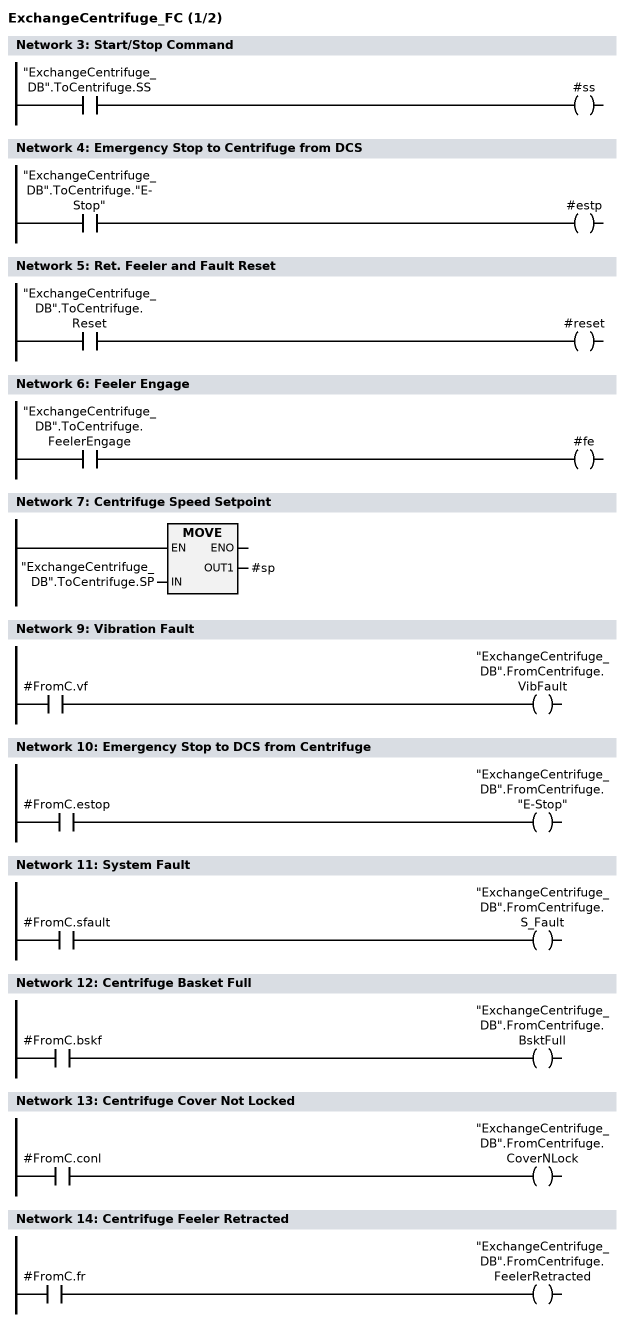
   RUNG wire#powerrail
      Contact( "ExchangeCentrifuge_DB".ToCentrifuge.SS )
      Coil( #ss )
   END_RUNG
   // the same network as SCL:
   #ss := "ExchangeCentrifuge_DB".ToCentrifuge.SS;
END_REGION

REGION Network 4: Emergency Stop to Centrifuge from DCS
   RUNG wire#powerrail
      Contact( "ExchangeCentrifuge_DB".ToCentrifuge."E-Stop" )
      Coil( #estp )
   END_RUNG
   // the same network as SCL:
   #estp := "ExchangeCentrifuge_DB".ToCentrifuge."E-Stop";
END_REGION

REGION Network 5: Ret. Feeler and Fault Reset
   RUNG wire#powerrail
      Contact( "ExchangeCentrifuge_DB".ToCentrifuge.Reset )
      Coil( #reset )
   END_RUNG
   // the same network as SCL:
   #reset := "ExchangeCentrifuge_DB".ToCentrifuge.Reset;
END_REGION

REGION Network 6: Feeler Engage
   RUNG wire#powerrail
      Contact( "ExchangeCentrifuge_DB".ToCentrifuge.FeelerEngage )
      Coil( #fe )
   END_RUNG
   // the same network as SCL:
   #fe := "ExchangeCentrifuge_DB".ToCentrifuge.FeelerEngage;
END_REGION

REGION Network 7: Centrifuge Speed Setpoint
   RUNG wire#powerrail
      Move(in := "ExchangeCentrifuge_DB".ToCentrifuge.SP, out1 => #sp)
   END_RUNG
   // the same network as SCL:
   #sp := "ExchangeCentrifuge_DB".ToCentrifuge.SP;
END_REGION

REGION Network 8: ////*********From Centrifuge to DCS**********////
   // Periphery Signal will be added to the contacts
END_REGION

REGION Network 9: Vibration Fault
   RUNG wire#powerrail
      Contact( #FromC.vf )
      Coil( "ExchangeCentrifuge_DB".FromCentrifuge.VibFault )
   END_RUNG
   // the same network as SCL:
   "ExchangeCentrifuge_DB".FromCentrifuge.VibFault := #FromC.vf;
END_REGION

REGION Network 10: Emergency Stop to DCS from Centrifuge
   RUNG wire#powerrail
      Contact( #FromC.estop )
      Coil( "ExchangeCentrifuge_DB".FromCentrifuge."E-Stop" )
   END_RUNG
   // the same network as SCL:
   "ExchangeCentrifuge_DB".FromCentrifuge."E-Stop" := #FromC.estop;
END_REGION

REGION Network 11: System Fault
   RUNG wire#powerrail
      Contact( #FromC.sfault )
      Coil( "ExchangeCentrifuge_DB".FromCentrifuge.S_Fault )
   END_RUNG
   // the same network as SCL:
   "ExchangeCentrifuge_DB".FromCentrifuge.S_Fault := #FromC.sfault;
END_REGION

REGION Network 12: Centrifuge Basket Full
   RUNG wire#powerrail
      Contact( #FromC.bskf )
      Coil( "ExchangeCentrifuge_DB".FromCentrifuge.BsktFull )
   END_RUNG
   // the same network as SCL:
   "ExchangeCentrifuge_DB".FromCentrifuge.BsktFull := #FromC.bskf;
END_REGION

REGION Network 13: Centrifuge Cover Not Locked
   RUNG wire#powerrail
      Contact( #FromC.conl )
      Coil( "ExchangeCentrifuge_DB".FromCentrifuge.CoverNLock )
   END_RUNG
   // the same network as SCL:
   "ExchangeCentrifuge_DB".FromCentrifuge.CoverNLock := #FromC.conl;
END_REGION

REGION Network 14: Centrifuge Feeler Retracted
   RUNG wire#powerrail
      Contact( #FromC.fr )
      Coil( "ExchangeCentrifuge_DB".FromCentrifuge.FeelerRetracted )
   END_RUNG
   // the same network as SCL:
   "ExchangeCentrifuge_DB".FromCentrifuge.FeelerRetracted := #FromC.fr;
END_REGION

REGION Network 15: Vibration Transmitter
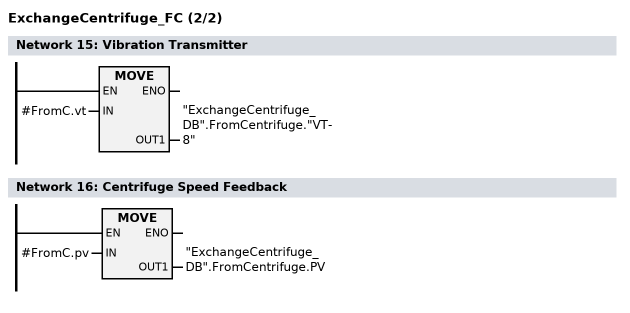
   RUNG wire#powerrail
      Move(in := #FromC.vt, out1 => "ExchangeCentrifuge_DB".FromCentrifuge."VT-8")
   END_RUNG
   // the same network as SCL:
   "ExchangeCentrifuge_DB".FromCentrifuge."VT-8" := #FromC.vt;
END_REGION

REGION Network 16: Centrifuge Speed Feedback
   RUNG wire#powerrail
      Move(in := #FromC.pv, out1 => "ExchangeCentrifuge_DB".FromCentrifuge.PV)
   END_RUNG
   // the same network as SCL:
   "ExchangeCentrifuge_DB".FromCentrifuge.PV := #FromC.pv;
END_REGION
END_FUNCTION

// folder: Outside Comms/ModBus Comms/CO/CO2/O2 R-401 Analizer

FUNCTION "Analizer_Modbus" : Void   // FC113, LAD
{ S7_Optimized_Access := 'TRUE' }
VERSION : 0.1
BEGIN

REGION Network 1: CO/CO2/O2 Analizer up to R-401 (Calcination)
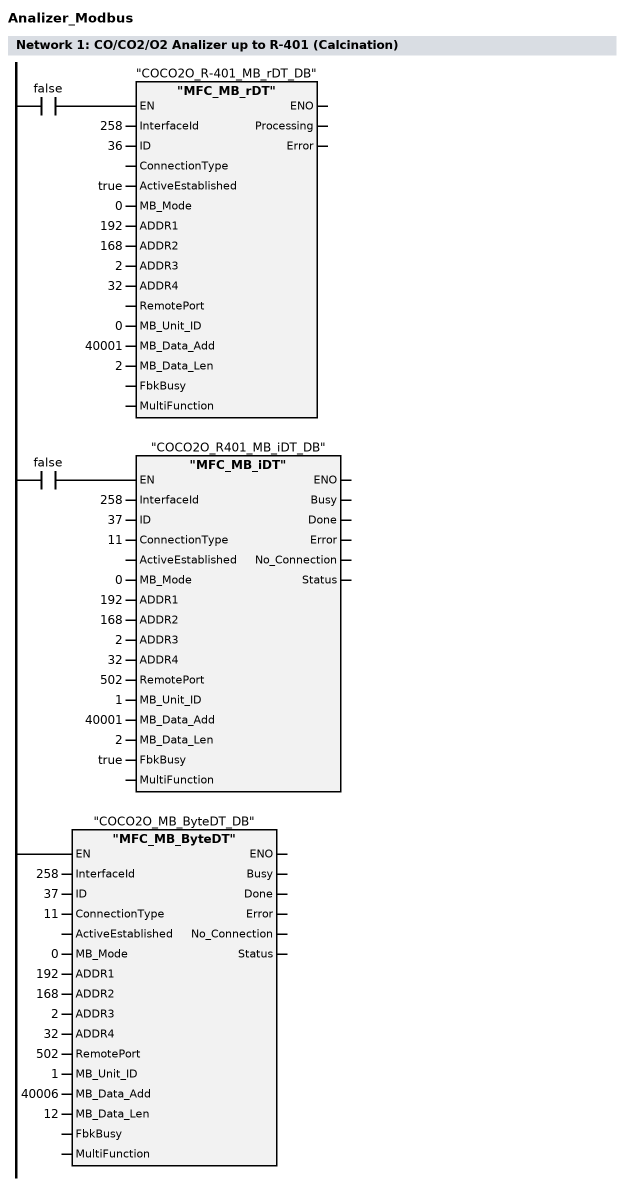
   RUNG wire#powerrail
      Contact( false )
      "COCO2O_R-401_MB_rDT_DB"(InterfaceId := 258, ID := 36, ConnectionType :=, ActiveEstablished := true, MB_Mode := 0, ADDR1 := 192, ADDR2 := 168, ADDR3 := 2, ADDR4 := 32, RemotePort :=, MB_Unit_ID := 0, MB_Data_Add := 40001, MB_Data_Len := 2, FbkBusy :=, MultiFunction :=, Processing =>, Error =>)
   END_RUNG
   RUNG wire#powerrail
      Contact( false )
      "COCO2O_R401_MB_iDT_DB"(InterfaceId := 258, ID := 37, ConnectionType := 11, ActiveEstablished :=, MB_Mode := 0, ADDR1 := 192, ADDR2 := 168, ADDR3 := 2, ADDR4 := 32, RemotePort := 502, MB_Unit_ID := 1, MB_Data_Add := 40001, MB_Data_Len := 2, FbkBusy := true, MultiFunction :=, Busy =>, Done =>, Error =>, No_Connection =>, Status =>)
   END_RUNG
   RUNG wire#powerrail
      "COCO2O_MB_ByteDT_DB"(InterfaceId := 258, ID := 37, ConnectionType := 11, ActiveEstablished :=, MB_Mode := 0, ADDR1 := 192, ADDR2 := 168, ADDR3 := 2, ADDR4 := 32, RemotePort := 502, MB_Unit_ID := 1, MB_Data_Add := 40006, MB_Data_Len := 12, FbkBusy :=, MultiFunction :=, Busy =>, Done =>, Error =>, No_Connection =>, Status =>)
   END_RUNG
   // the same network as SCL:
   IF false THEN
       "COCO2O_R-401_MB_rDT_DB"(InterfaceId := 258,   // "MFC_MB_rDT"
                               ID := 36,
                               ActiveEstablished := true,
                               MB_Mode := 0,
                               ADDR1 := 192,
                               ADDR2 := 168,
                               ADDR3 := 2,
                               ADDR4 := 32,
                               MB_Unit_ID := 0,
                               MB_Data_Add := 40001,
                               MB_Data_Len := 2);
       "COCO2O_R401_MB_iDT_DB"(InterfaceId := 258,   // "MFC_MB_iDT"
                               ID := 37,
                               ConnectionType := 11,
                               MB_Mode := 0,
                               ADDR1 := 192,
                               ADDR2 := 168,
                               ADDR3 := 2,
                               ADDR4 := 32,
                               RemotePort := 502,
                               MB_Unit_ID := 1,
                               MB_Data_Add := 40001,
                               MB_Data_Len := 2,
                               FbkBusy := true);
   END_IF;
   "COCO2O_MB_ByteDT_DB"(InterfaceId := 258,   // "MFC_MB_ByteDT"
                         ID := 37,
                         ConnectionType := 11,
                         MB_Mode := 0,
                         ADDR1 := 192,
                         ADDR2 := 168,
                         ADDR3 := 2,
                         ADDR4 := 32,
                         RemotePort := 502,
                         MB_Unit_ID := 1,
                         MB_Data_Add := 40006,
                         MB_Data_Len := 12);
END_REGION
END_FUNCTION

// folder: Outside Comms/ModBus Comms/EurothermControllers

FUNCTION_BLOCK "Eurotherm_MB_FB"   // FB29, LAD
TITLE = Modbus Block for Real Data Type
{ S7_Optimized_Access := 'TRUE' }
AUTHOR : JL
VERSION : 0.1
   VAR_INPUT
      InterfaceId : Hw_Any;   // HW-identifier of IE-interface submodule
      ID : Conn_Ouc;   // connection reference / identifier
      ConnectionType : Byte;   // type of connection: 11=TCP/IP, 19=UDP (17=TCP/IP)
      ActiveEstablished : Bool := true;   // active/passive connection establishment
      Disconnect : Bool;
      MB_Mode : Byte;
      ADDR1 : Byte;   // IPv4 address
      ADDR2 : Byte;   // IPv4 address
      ADDR3 : Byte;   // IPv4 address
      ADDR4 : Byte;   // IPv4 address
      RemotePort : UInt;   // remote UDP/TCP port number
      MB_Unit_ID : Byte;   // The Modbus slave address
      MB_Data_Add : UDInt;   // Modbus Data Address
      MB_Data_Len : UInt;   // Modbus Data Length
      ManualTrigger : Bool;
      MultiFunction : Bool;   // Depend of the status of the other calls same MB
   END_VAR
   VAR_OUTPUT
      Processing : Bool;
      Done : Bool;
      Busy : Bool;
      Error : Bool;
      ErrorStatus : Word;
   END_VAR
   VAR
      MB_CLIENT_Instance : MB_CLIENT;
      MB_Ctrl : Struct
         REQ : Bool;
         REQ_Again : Bool;
         Disconnect : Bool := false;
         MB_Mode : Byte;   // Modbus Mode
         MB_Data_Address : UDInt;   // Modbus Data Address
         MB_Data_Length : UInt;   // Modbus Data Length
         Connect : TCON_IP_v4;   // Connect Parameters Client
      END_STRUCT;
      MB_Data : Struct
         Buffer : Array[1..16] of Int;
      END_STRUCT;
      "Timer" : Struct
         "1" : IEC_TIMER;
         "2" : IEC_TIMER;
      END_STRUCT;
      OS : Struct
         bit : Array[0..31] of Bool;
      END_STRUCT;
      Process : Struct
         Start : Bool;
         CmdRead : Bool;
         End : Bool;
      END_STRUCT;
   END_VAR
   VAR_TEMP   // added for the SCL form of the ladder/FBD networks
      _w1 : Bool;
      _w2 : Bool;
      _w3 : Bool;
   END_VAR
   // MB_Ctrl.Connect.InterfaceId := 258;
   // MB_Ctrl.Connect.ID := 11;
   // MB_Ctrl.Connect.ConnectionType := 11;
   // MB_Ctrl.Connect.ActiveEstablished := 1;
   // MB_Ctrl.Connect.RemoteAddress.ADDR[1] := 192;
   // MB_Ctrl.Connect.RemoteAddress.ADDR[2] := 168;
   // MB_Ctrl.Connect.RemoteAddress.ADDR[3] := 2;
   // MB_Ctrl.Connect.RemoteAddress.ADDR[4] := 11;
   // MB_Ctrl.Connect.RemotePort := 502;
BEGIN

REGION Network 1 (SCL): Block Parameters
   #MB_Ctrl.Connect.InterfaceId := #InterfaceId;
   #MB_Ctrl.Connect.ID := #ID;
   #MB_Ctrl.Connect.ConnectionType:=#ConnectionType;
   #MB_Ctrl.Disconnect := #Disconnect;
   #MB_Ctrl.MB_Mode:=#MB_Mode;
   #MB_Ctrl.Connect.ActiveEstablished:=#ActiveEstablished;
   #MB_Ctrl.Connect.RemoteAddress.ADDR[1] := #ADDR1;
   #MB_Ctrl.Connect.RemoteAddress.ADDR[2] := #ADDR2;
   #MB_Ctrl.Connect.RemoteAddress.ADDR[3] := #ADDR3;
   #MB_Ctrl.Connect.RemoteAddress.ADDR[4] := #ADDR4;
   #MB_Ctrl.Connect.RemotePort := #RemotePort;
   #MB_CLIENT_Instance.MB_Unit_ID := #MB_Unit_ID;
   #MB_Ctrl.MB_Data_Address := #MB_Data_Add;
   #MB_Ctrl.MB_Data_Length := #MB_Data_Len;
   //#MB_Ctrl.Disconnect := #FbkBusy;
END_REGION

REGION Network 2: Reading Indication
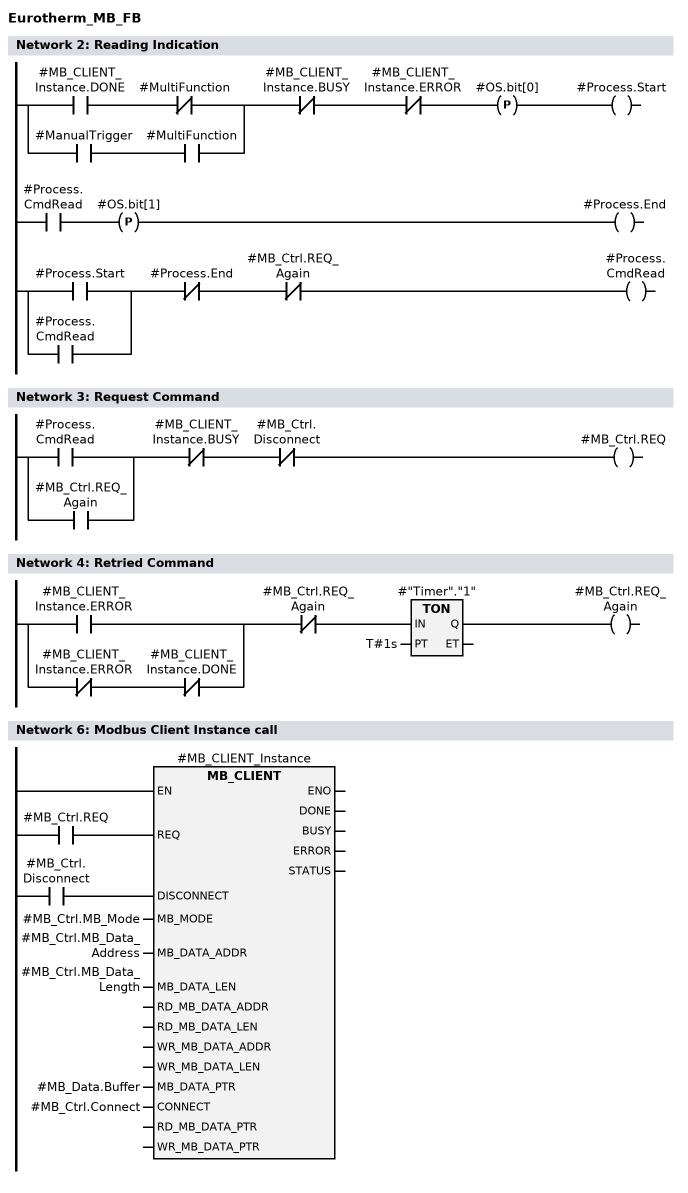
   RUNG wire#powerrail
      Contact( #MB_CLIENT_Instance.DONE )
      I_Contact( #MultiFunction )
      wire#w1
      I_Contact( #MB_CLIENT_Instance.BUSY )
      I_Contact( #MB_CLIENT_Instance.ERROR )
      P_Trig( #OS.bit[0] )
      Coil( #Process.Start )
   END_RUNG
   RUNG wire#powerrail
      Contact( #ManualTrigger )
      Contact( #MultiFunction )
   END_RUNG wire#w1
   RUNG wire#powerrail
      Contact( #Process.CmdRead )
      P_Trig( #OS.bit[1] )
      Coil( #Process.End )
   END_RUNG
   RUNG wire#powerrail
      Contact( #Process.Start )
      wire#w2
      I_Contact( #Process.End )
      I_Contact( #MB_Ctrl.REQ_Again )
      Coil( #Process.CmdRead )
   END_RUNG
   RUNG wire#powerrail
      Contact( #Process.CmdRead )
   END_RUNG wire#w2
   // the same network as SCL:
   #_w1 := ((#MB_CLIENT_Instance.DONE AND NOT #MultiFunction) OR (#ManualTrigger AND #MultiFunction)) AND NOT #MB_CLIENT_Instance.BUSY AND NOT #MB_CLIENT_Instance.ERROR;
   #_w2 := #_w1 AND NOT #OS.bit[0];   // rising edge
   #OS.bit[0] := #_w1;
   #Process.Start := #_w2;
   #_w3 := #Process.CmdRead AND NOT #OS.bit[1];   // rising edge
   #OS.bit[1] := #Process.CmdRead;
   #Process.End := #_w3;
   #Process.CmdRead := (#Process.Start OR #Process.CmdRead) AND NOT #Process.End AND NOT #MB_Ctrl.REQ_Again;
END_REGION

REGION Network 3: Request Command
   RUNG wire#powerrail
      Contact( #Process.CmdRead )
      wire#w1
      I_Contact( #MB_CLIENT_Instance.BUSY )
      I_Contact( #MB_Ctrl.Disconnect )
      Coil( #MB_Ctrl.REQ )
   END_RUNG
   RUNG wire#powerrail
      Contact( #MB_Ctrl.REQ_Again )
   END_RUNG wire#w1
   // the same network as SCL:
   #MB_Ctrl.REQ := (#Process.CmdRead OR #MB_Ctrl.REQ_Again) AND NOT #MB_CLIENT_Instance.BUSY AND NOT #MB_Ctrl.Disconnect;
END_REGION

REGION Network 4: Retried Command
   #"Timer"."1".TON(IN := (#MB_CLIENT_Instance.ERROR OR (NOT #MB_CLIENT_Instance.ERROR AND NOT #MB_CLIENT_Instance.DONE)) AND NOT #MB_Ctrl.REQ_Again,
                    PT := T#1s);
   #MB_Ctrl.REQ_Again := #"Timer"."1".Q;
END_REGION

REGION Network 5 (SCL)
   IF #MB_CLIENT_Instance.ERROR AND #Timer."1".Q THEN
       #MB_CLIENT_Instance.Connected := TRUE;
   END_IF;
END_REGION

REGION Network 6: Modbus Client Instance call
   #MB_CLIENT_Instance(REQ := #MB_Ctrl.REQ,   // MB_CLIENT
                       DISCONNECT := #MB_Ctrl.Disconnect,
                       MB_MODE := #MB_Ctrl.MB_Mode,
                       MB_DATA_ADDR := #MB_Ctrl.MB_Data_Address,
                       MB_DATA_LEN := #MB_Ctrl.MB_Data_Length,
                       MB_DATA_PTR := #MB_Data.Buffer,
                       CONNECT := #MB_Ctrl.Connect);
END_REGION

REGION Network 7 (SCL)
   #Processing := #MB_CLIENT_Instance.BUSY AND NOT #MB_CLIENT_Instance.DONE;
   #Done := #MB_CLIENT_Instance.DONE AND NOT #MB_CLIENT_Instance.BUSY AND NOT #MB_CLIENT_Instance.ERROR;
   #Busy := #MB_CLIENT_Instance.BUSY AND NOT #MB_CLIENT_Instance.DONE;
   #Error := #MB_CLIENT_Instance.ERROR;
   #ErrorStatus := #MB_CLIENT_Instance.STATUS;
END_REGION
END_FUNCTION_BLOCK

FUNCTION "AddrMoves" : Void   // FC97, SCL
{ S7_Optimized_Access := 'TRUE' }
VERSION : 0.1
   VAR_INPUT
      StartAddr : UDInt;
      EndAddr : UDInt;
      NextAddr : Bool;
      Initialize : Bool;
   END_VAR
   VAR_IN_OUT
      CurrentAddr : UDInt;
      Down : Bool;
      UP : Bool;
      RisingUp : Bool;
   END_VAR
BEGIN
   //********bbbbbbbbbbbbbbbbbbbb/////////////////
   IF #StartAddr > 0 AND #EndAddr > #StartAddr AND NOT #Initialize THEN

       IF NOT #NextAddr THEN   //Input is at Zero
           #Down := True;
       END_IF;

       IF  #NextAddr THEN      //Input is at One
           #UP := True;
       END_IF;

       IF #Down AND #NextAddr THEN     //Detection of the Rising edge 
           #Down := false;
           #RisingUp := TRUE;
       ELSE
           #RisingUp := FALSE;
       END_IF;




       IF   #RisingUp  THEN //Rise adge detected
           IF  #CurrentAddr < #EndAddr THEN
               #CurrentAddr := #CurrentAddr + 1;

           ELSE
               #CurrentAddr := #StartAddr;
           END_IF;

       END_IF;

   ELSE         //To initialize the actual address
       #CurrentAddr := #StartAddr;
       #Down := FALSE;
       #UP := FALSE;
       #RisingUp := FALSE;

   END_IF;
END_FUNCTION

// folder: Outside Comms/ModBus Comms/EurothermControllers/TC-4011A

FUNCTION "TC_4011A" : Void   // FC31, LAD
{ S7_Optimized_Access := 'TRUE' }
VERSION : 0.1
   VAR_TEMP
      MBAddress : UDInt;
      Run : Bool;
      Reset : Bool;
      notProcess : Bool;
   END_VAR
BEGIN

REGION Network 1 (SCL)
   //Data Read 1
   //MOVE_BLK(IN := "Eurothem_Data".Read.Read1.Slaves.Slave1[1],
      //      COUNT := 12,
       //     OUT => "TC-4011A_R1".MB_Data.Buffer[1]);
END_REGION

REGION Network 2: Read Data 1
   // R1=30001
   // R2=31280
   // R3=30023
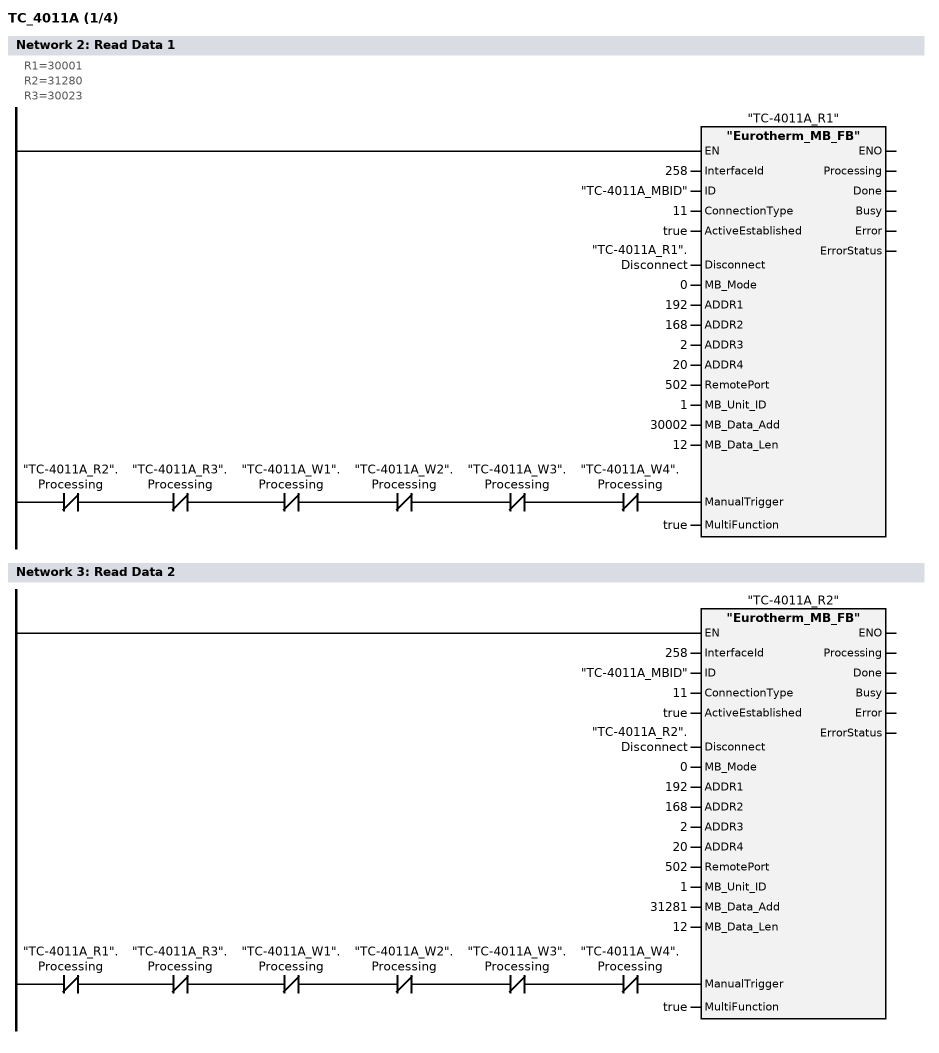
   RUNG wire#powerrail
      "TC-4011A_R1"(ManualTrigger := wire#w1, InterfaceId := 258, ID := "TC-4011A_MBID", ConnectionType := 11, ActiveEstablished := true, Disconnect := "TC-4011A_R1".Disconnect, MB_Mode := 0, ADDR1 := 192, ADDR2 := 168, ADDR3 := 2, ADDR4 := 20, RemotePort := 502, MB_Unit_ID := 1, MB_Data_Add := 30002, MB_Data_Len := 12, MultiFunction := true, Processing =>, Done =>, Busy =>, Error =>, ErrorStatus =>)
   END_RUNG
   RUNG wire#powerrail
      I_Contact( "TC-4011A_R2".Processing )
      I_Contact( "TC-4011A_R3".Processing )
      I_Contact( "TC-4011A_W1".Processing )
      I_Contact( "TC-4011A_W2".Processing )
      I_Contact( "TC-4011A_W3".Processing )
      I_Contact( "TC-4011A_W4".Processing )
   END_RUNG wire#w1
   // the same network as SCL:
   "TC-4011A_R1"(InterfaceId := 258,   // "Eurotherm_MB_FB"
                 ID := "TC-4011A_MBID",
                 ConnectionType := 11,
                 ActiveEstablished := true,
                 Disconnect := "TC-4011A_R1".Disconnect,
                 MB_Mode := 0,
                 ADDR1 := 192,
                 ADDR2 := 168,
                 ADDR3 := 2,
                 ADDR4 := 20,
                 RemotePort := 502,
                 MB_Unit_ID := 1,
                 MB_Data_Add := 30002,
                 MB_Data_Len := 12,
                 ManualTrigger := NOT "TC-4011A_R2".Processing AND NOT "TC-4011A_R3".Processing AND NOT "TC-4011A_W1".Processing AND NOT "TC-4011A_W2".Processing AND NOT "TC-4011A_W3".Processing AND NOT "TC-4011A_W4".Processing,
                 MultiFunction := true);
END_REGION

REGION Network 3: Read Data 2
   RUNG wire#powerrail
      "TC-4011A_R2"(ManualTrigger := wire#w1, InterfaceId := 258, ID := "TC-4011A_MBID", ConnectionType := 11, ActiveEstablished := true, Disconnect := "TC-4011A_R2".Disconnect, MB_Mode := 0, ADDR1 := 192, ADDR2 := 168, ADDR3 := 2, ADDR4 := 20, RemotePort := 502, MB_Unit_ID := 1, MB_Data_Add := 31281, MB_Data_Len := 12, MultiFunction := true, Processing =>, Done =>, Busy =>, Error =>, ErrorStatus =>)
   END_RUNG
   RUNG wire#powerrail
      I_Contact( "TC-4011A_R1".Processing )
      I_Contact( "TC-4011A_R3".Processing )
      I_Contact( "TC-4011A_W1".Processing )
      I_Contact( "TC-4011A_W2".Processing )
      I_Contact( "TC-4011A_W3".Processing )
      I_Contact( "TC-4011A_W4".Processing )
   END_RUNG wire#w1
   // the same network as SCL:
   "TC-4011A_R2"(InterfaceId := 258,   // "Eurotherm_MB_FB"
                 ID := "TC-4011A_MBID",
                 ConnectionType := 11,
                 ActiveEstablished := true,
                 Disconnect := "TC-4011A_R2".Disconnect,
                 MB_Mode := 0,
                 ADDR1 := 192,
                 ADDR2 := 168,
                 ADDR3 := 2,
                 ADDR4 := 20,
                 RemotePort := 502,
                 MB_Unit_ID := 1,
                 MB_Data_Add := 31281,
                 MB_Data_Len := 12,
                 ManualTrigger := NOT "TC-4011A_R1".Processing AND NOT "TC-4011A_R3".Processing AND NOT "TC-4011A_W1".Processing AND NOT "TC-4011A_W2".Processing AND NOT "TC-4011A_W3".Processing AND NOT "TC-4011A_W4".Processing,
                 MultiFunction := true);
END_REGION

REGION Network 4: Read Data 3
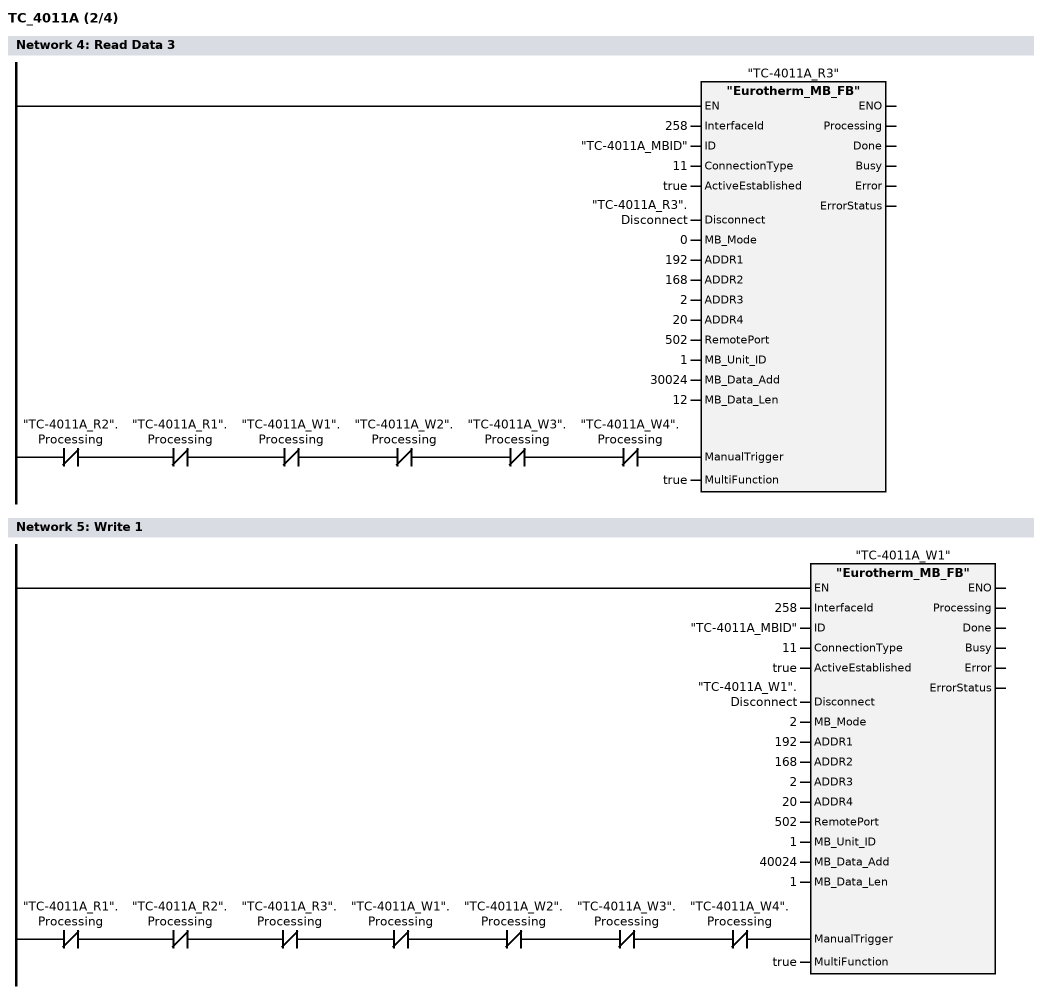
   RUNG wire#powerrail
      "TC-4011A_R3"(ManualTrigger := wire#w1, InterfaceId := 258, ID := "TC-4011A_MBID", ConnectionType := 11, ActiveEstablished := true, Disconnect := "TC-4011A_R3".Disconnect, MB_Mode := 0, ADDR1 := 192, ADDR2 := 168, ADDR3 := 2, ADDR4 := 20, RemotePort := 502, MB_Unit_ID := 1, MB_Data_Add := 30024, MB_Data_Len := 12, MultiFunction := true, Processing =>, Done =>, Busy =>, Error =>, ErrorStatus =>)
   END_RUNG
   RUNG wire#powerrail
      I_Contact( "TC-4011A_R2".Processing )
      I_Contact( "TC-4011A_R1".Processing )
      I_Contact( "TC-4011A_W1".Processing )
      I_Contact( "TC-4011A_W2".Processing )
      I_Contact( "TC-4011A_W3".Processing )
      I_Contact( "TC-4011A_W4".Processing )
   END_RUNG wire#w1
   // the same network as SCL:
   "TC-4011A_R3"(InterfaceId := 258,   // "Eurotherm_MB_FB"
                 ID := "TC-4011A_MBID",
                 ConnectionType := 11,
                 ActiveEstablished := true,
                 Disconnect := "TC-4011A_R3".Disconnect,
                 MB_Mode := 0,
                 ADDR1 := 192,
                 ADDR2 := 168,
                 ADDR3 := 2,
                 ADDR4 := 20,
                 RemotePort := 502,
                 MB_Unit_ID := 1,
                 MB_Data_Add := 30024,
                 MB_Data_Len := 12,
                 ManualTrigger := NOT "TC-4011A_R2".Processing AND NOT "TC-4011A_R1".Processing AND NOT "TC-4011A_W1".Processing AND NOT "TC-4011A_W2".Processing AND NOT "TC-4011A_W3".Processing AND NOT "TC-4011A_W4".Processing,
                 MultiFunction := true);
END_REGION

REGION Network 5: Write 1
   RUNG wire#powerrail
      "TC-4011A_W1"(ManualTrigger := wire#w1, InterfaceId := 258, ID := "TC-4011A_MBID", ConnectionType := 11, ActiveEstablished := true, Disconnect := "TC-4011A_W1".Disconnect, MB_Mode := 2, ADDR1 := 192, ADDR2 := 168, ADDR3 := 2, ADDR4 := 20, RemotePort := 502, MB_Unit_ID := 1, MB_Data_Add := 40024, MB_Data_Len := 1, MultiFunction := true, Processing =>, Done =>, Busy =>, Error =>, ErrorStatus =>)
   END_RUNG
   RUNG wire#powerrail
      I_Contact( "TC-4011A_R1".Processing )
      I_Contact( "TC-4011A_R2".Processing )
      I_Contact( "TC-4011A_R3".Processing )
      I_Contact( "TC-4011A_W1".Processing )
      I_Contact( "TC-4011A_W2".Processing )
      I_Contact( "TC-4011A_W3".Processing )
      I_Contact( "TC-4011A_W4".Processing )
   END_RUNG wire#w1
   // the same network as SCL:
   "TC-4011A_W1"(InterfaceId := 258,   // "Eurotherm_MB_FB"
                 ID := "TC-4011A_MBID",
                 ConnectionType := 11,
                 ActiveEstablished := true,
                 Disconnect := "TC-4011A_W1".Disconnect,
                 MB_Mode := 2,
                 ADDR1 := 192,
                 ADDR2 := 168,
                 ADDR3 := 2,
                 ADDR4 := 20,
                 RemotePort := 502,
                 MB_Unit_ID := 1,
                 MB_Data_Add := 40024,
                 MB_Data_Len := 1,
                 ManualTrigger := NOT "TC-4011A_R1".Processing AND NOT "TC-4011A_R2".Processing AND NOT "TC-4011A_R3".Processing AND NOT "TC-4011A_W1".Processing AND NOT "TC-4011A_W2".Processing AND NOT "TC-4011A_W3".Processing AND NOT "TC-4011A_W4".Processing,
                 MultiFunction := true);
END_REGION

REGION Network 6: Write 2
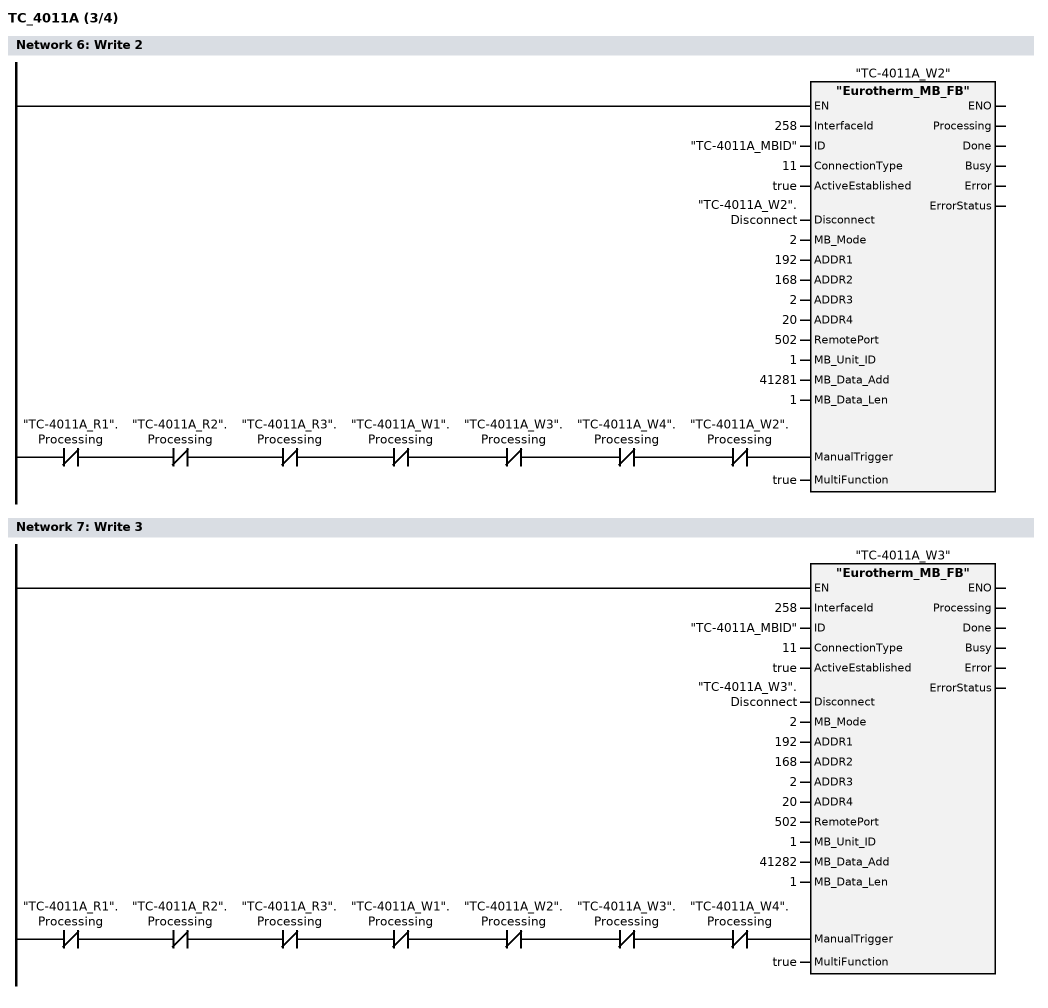
   RUNG wire#powerrail
      "TC-4011A_W2"(ManualTrigger := wire#w1, InterfaceId := 258, ID := "TC-4011A_MBID", ConnectionType := 11, ActiveEstablished := true, Disconnect := "TC-4011A_W2".Disconnect, MB_Mode := 2, ADDR1 := 192, ADDR2 := 168, ADDR3 := 2, ADDR4 := 20, RemotePort := 502, MB_Unit_ID := 1, MB_Data_Add := 41281, MB_Data_Len := 1, MultiFunction := true, Processing =>, Done =>, Busy =>, Error =>, ErrorStatus =>)
   END_RUNG
   RUNG wire#powerrail
      I_Contact( "TC-4011A_R1".Processing )
      I_Contact( "TC-4011A_R2".Processing )
      I_Contact( "TC-4011A_R3".Processing )
      I_Contact( "TC-4011A_W1".Processing )
      I_Contact( "TC-4011A_W3".Processing )
      I_Contact( "TC-4011A_W4".Processing )
      I_Contact( "TC-4011A_W2".Processing )
   END_RUNG wire#w1
   // the same network as SCL:
   "TC-4011A_W2"(InterfaceId := 258,   // "Eurotherm_MB_FB"
                 ID := "TC-4011A_MBID",
                 ConnectionType := 11,
                 ActiveEstablished := true,
                 Disconnect := "TC-4011A_W2".Disconnect,
                 MB_Mode := 2,
                 ADDR1 := 192,
                 ADDR2 := 168,
                 ADDR3 := 2,
                 ADDR4 := 20,
                 RemotePort := 502,
                 MB_Unit_ID := 1,
                 MB_Data_Add := 41281,
                 MB_Data_Len := 1,
                 ManualTrigger := NOT "TC-4011A_R1".Processing AND NOT "TC-4011A_R2".Processing AND NOT "TC-4011A_R3".Processing AND NOT "TC-4011A_W1".Processing AND NOT "TC-4011A_W3".Processing AND NOT "TC-4011A_W4".Processing AND NOT "TC-4011A_W2".Processing,
                 MultiFunction := true);
END_REGION

REGION Network 7: Write 3
   RUNG wire#powerrail
      "TC-4011A_W3"(ManualTrigger := wire#w1, InterfaceId := 258, ID := "TC-4011A_MBID", ConnectionType := 11, ActiveEstablished := true, Disconnect := "TC-4011A_W3".Disconnect, MB_Mode := 2, ADDR1 := 192, ADDR2 := 168, ADDR3 := 2, ADDR4 := 20, RemotePort := 502, MB_Unit_ID := 1, MB_Data_Add := 41282, MB_Data_Len := 1, MultiFunction := true, Processing =>, Done =>, Busy =>, Error =>, ErrorStatus =>)
   END_RUNG
   RUNG wire#powerrail
      I_Contact( "TC-4011A_R1".Processing )
      I_Contact( "TC-4011A_R2".Processing )
      I_Contact( "TC-4011A_R3".Processing )
      I_Contact( "TC-4011A_W1".Processing )
      I_Contact( "TC-4011A_W2".Processing )
      I_Contact( "TC-4011A_W3".Processing )
      I_Contact( "TC-4011A_W4".Processing )
   END_RUNG wire#w1
   // the same network as SCL:
   "TC-4011A_W3"(InterfaceId := 258,   // "Eurotherm_MB_FB"
                 ID := "TC-4011A_MBID",
                 ConnectionType := 11,
                 ActiveEstablished := true,
                 Disconnect := "TC-4011A_W3".Disconnect,
                 MB_Mode := 2,
                 ADDR1 := 192,
                 ADDR2 := 168,
                 ADDR3 := 2,
                 ADDR4 := 20,
                 RemotePort := 502,
                 MB_Unit_ID := 1,
                 MB_Data_Add := 41282,
                 MB_Data_Len := 1,
                 ManualTrigger := NOT "TC-4011A_R1".Processing AND NOT "TC-4011A_R2".Processing AND NOT "TC-4011A_R3".Processing AND NOT "TC-4011A_W1".Processing AND NOT "TC-4011A_W2".Processing AND NOT "TC-4011A_W3".Processing AND NOT "TC-4011A_W4".Processing,
                 MultiFunction := true);
END_REGION

REGION Network 8: Write 4
